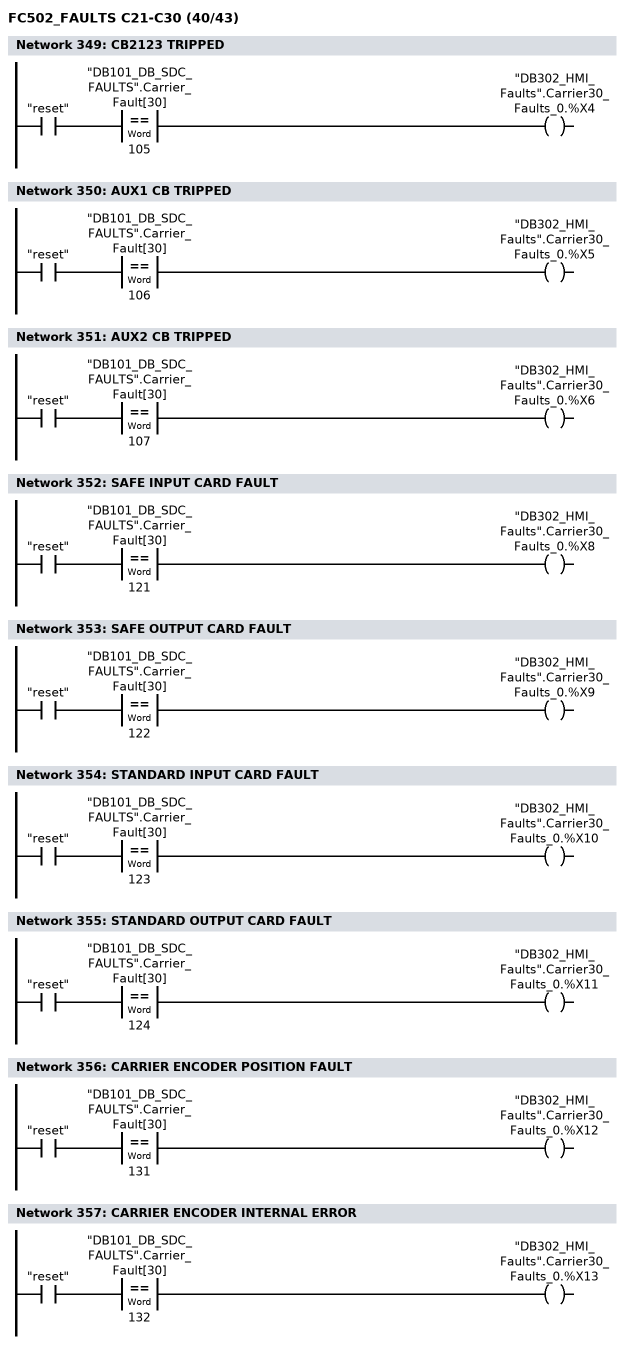
   RUNG wire#powerrail
      Contact( "reset" )
      { S7_Templates := "SrcType := Word" } EQ_Contact(in1 := "DB101_DB_SDC_FAULTS".Carrier_Fault[30], in2 := 105)
      Coil( "DB302_HMI_Faults".Carrier30_Faults_0.%X4 )
   END_RUNG
   // the same network as SCL:
   "DB302_HMI_Faults".Carrier30_Faults_0.%X4 := "reset" AND ("DB101_DB_SDC_FAULTS".Carrier_Fault[30] = 105);
END_REGION

REGION Network 350: AUX1 CB TRIPPED
   RUNG wire#powerrail
      Contact( "reset" )
      { S7_Templates := "SrcType := Word" } EQ_Contact(in1 := "DB101_DB_SDC_FAULTS".Carrier_Fault[30], in2 := 106)
      Coil( "DB302_HMI_Faults".Carrier30_Faults_0.%X5 )
   END_RUNG
   // the same network as SCL:
   "DB302_HMI_Faults".Carrier30_Faults_0.%X5 := "reset" AND ("DB101_DB_SDC_FAULTS".Carrier_Fault[30] = 106);
END_REGION

REGION Network 351: AUX2 CB TRIPPED
   RUNG wire#powerrail
      Contact( "reset" )
      { S7_Templates := "SrcType := Word" } EQ_Contact(in1 := "DB101_DB_SDC_FAULTS".Carrier_Fault[30], in2 := 107)
      Coil( "DB302_HMI_Faults".Carrier30_Faults_0.%X6 )
   END_RUNG
   // the same network as SCL:
   "DB302_HMI_Faults".Carrier30_Faults_0.%X6 := "reset" AND ("DB101_DB_SDC_FAULTS".Carrier_Fault[30] = 107);
END_REGION

REGION Network 352: SAFE INPUT CARD FAULT
   RUNG wire#powerrail
      Contact( "reset" )
      { S7_Templates := "SrcType := Word" } EQ_Contact(in1 := "DB101_DB_SDC_FAULTS".Carrier_Fault[30], in2 := 121)
      Coil( "DB302_HMI_Faults".Carrier30_Faults_0.%X8 )
   END_RUNG
   // the same network as SCL:
   "DB302_HMI_Faults".Carrier30_Faults_0.%X8 := "reset" AND ("DB101_DB_SDC_FAULTS".Carrier_Fault[30] = 121);
END_REGION

REGION Network 353: SAFE OUTPUT CARD FAULT
   RUNG wire#powerrail
      Contact( "reset" )
      { S7_Templates := "SrcType := Word" } EQ_Contact(in1 := "DB101_DB_SDC_FAULTS".Carrier_Fault[30], in2 := 122)
      Coil( "DB302_HMI_Faults".Carrier30_Faults_0.%X9 )
   END_RUNG
   // the same network as SCL:
   "DB302_HMI_Faults".Carrier30_Faults_0.%X9 := "reset" AND ("DB101_DB_SDC_FAULTS".Carrier_Fault[30] = 122);
END_REGION

REGION Network 354: STANDARD INPUT CARD FAULT
   RUNG wire#powerrail
      Contact( "reset" )
      { S7_Templates := "SrcType := Word" } EQ_Contact(in1 := "DB101_DB_SDC_FAULTS".Carrier_Fault[30], in2 := 123)
      Coil( "DB302_HMI_Faults".Carrier30_Faults_0.%X10 )
   END_RUNG
   // the same network as SCL:
   "DB302_HMI_Faults".Carrier30_Faults_0.%X10 := "reset" AND ("DB101_DB_SDC_FAULTS".Carrier_Fault[30] = 123);
END_REGION

REGION Network 355: STANDARD OUTPUT CARD FAULT
   RUNG wire#powerrail
      Contact( "reset" )
      { S7_Templates := "SrcType := Word" } EQ_Contact(in1 := "DB101_DB_SDC_FAULTS".Carrier_Fault[30], in2 := 124)
      Coil( "DB302_HMI_Faults".Carrier30_Faults_0.%X11 )
   END_RUNG
   // the same network as SCL:
   "DB302_HMI_Faults".Carrier30_Faults_0.%X11 := "reset" AND ("DB101_DB_SDC_FAULTS".Carrier_Fault[30] = 124);
END_REGION

REGION Network 356: CARRIER ENCODER POSITION FAULT
   RUNG wire#powerrail
      Contact( "reset" )
      { S7_Templates := "SrcType := Word" } EQ_Contact(in1 := "DB101_DB_SDC_FAULTS".Carrier_Fault[30], in2 := 131)
      Coil( "DB302_HMI_Faults".Carrier30_Faults_0.%X12 )
   END_RUNG
   // the same network as SCL:
   "DB302_HMI_Faults".Carrier30_Faults_0.%X12 := "reset" AND ("DB101_DB_SDC_FAULTS".Carrier_Fault[30] = 131);
END_REGION

REGION Network 357: CARRIER ENCODER INTERNAL ERROR
   RUNG wire#powerrail
      Contact( "reset" )
      { S7_Templates := "SrcType := Word" } EQ_Contact(in1 := "DB101_DB_SDC_FAULTS".Carrier_Fault[30], in2 := 132)
      Coil( "DB302_HMI_Faults".Carrier30_Faults_0.%X13 )
   END_RUNG
   // the same network as SCL:
   "DB302_HMI_Faults".Carrier30_Faults_0.%X13 := "reset" AND ("DB101_DB_SDC_FAULTS".Carrier_Fault[30] = 132);
END_REGION

REGION Network 358: CARRIER ENCODER COMM FAULT
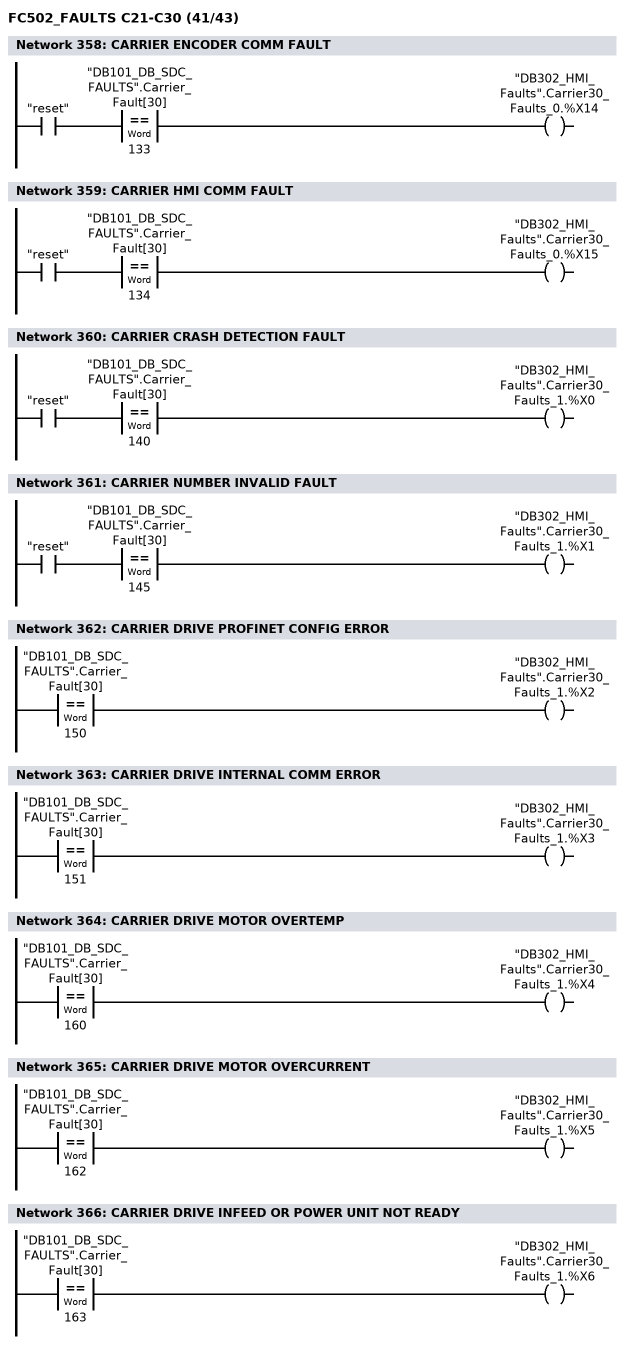
   RUNG wire#powerrail
      Contact( "reset" )
      { S7_Templates := "SrcType := Word" } EQ_Contact(in1 := "DB101_DB_SDC_FAULTS".Carrier_Fault[30], in2 := 133)
      Coil( "DB302_HMI_Faults".Carrier30_Faults_0.%X14 )
   END_RUNG
   // the same network as SCL:
   "DB302_HMI_Faults".Carrier30_Faults_0.%X14 := "reset" AND ("DB101_DB_SDC_FAULTS".Carrier_Fault[30] = 133);
END_REGION

REGION Network 359: CARRIER HMI COMM FAULT
   RUNG wire#powerrail
      Contact( "reset" )
      { S7_Templates := "SrcType := Word" } EQ_Contact(in1 := "DB101_DB_SDC_FAULTS".Carrier_Fault[30], in2 := 134)
      Coil( "DB302_HMI_Faults".Carrier30_Faults_0.%X15 )
   END_RUNG
   // the same network as SCL:
   "DB302_HMI_Faults".Carrier30_Faults_0.%X15 := "reset" AND ("DB101_DB_SDC_FAULTS".Carrier_Fault[30] = 134);
END_REGION

REGION Network 360: CARRIER CRASH DETECTION FAULT
   RUNG wire#powerrail
      Contact( "reset" )
      { S7_Templates := "SrcType := Word" } EQ_Contact(in1 := "DB101_DB_SDC_FAULTS".Carrier_Fault[30], in2 := 140)
      Coil( "DB302_HMI_Faults".Carrier30_Faults_1.%X0 )
   END_RUNG
   // the same network as SCL:
   "DB302_HMI_Faults".Carrier30_Faults_1.%X0 := "reset" AND ("DB101_DB_SDC_FAULTS".Carrier_Fault[30] = 140);
END_REGION

REGION Network 361: CARRIER NUMBER INVALID FAULT
   RUNG wire#powerrail
      Contact( "reset" )
      { S7_Templates := "SrcType := Word" } EQ_Contact(in1 := "DB101_DB_SDC_FAULTS".Carrier_Fault[30], in2 := 145)
      Coil( "DB302_HMI_Faults".Carrier30_Faults_1.%X1 )
   END_RUNG
   // the same network as SCL:
   "DB302_HMI_Faults".Carrier30_Faults_1.%X1 := "reset" AND ("DB101_DB_SDC_FAULTS".Carrier_Fault[30] = 145);
END_REGION

REGION Network 362: CARRIER DRIVE PROFINET CONFIG ERROR
   RUNG wire#powerrail
      { S7_Templates := "SrcType := Word" } EQ_Contact(in1 := "DB101_DB_SDC_FAULTS".Carrier_Fault[30], in2 := 150)
      Coil( "DB302_HMI_Faults".Carrier30_Faults_1.%X2 )
   END_RUNG
   // the same network as SCL:
   "DB302_HMI_Faults".Carrier30_Faults_1.%X2 := "DB101_DB_SDC_FAULTS".Carrier_Fault[30] = 150;
END_REGION

REGION Network 363: CARRIER DRIVE INTERNAL COMM ERROR
   RUNG wire#powerrail
      { S7_Templates := "SrcType := Word" } EQ_Contact(in1 := "DB101_DB_SDC_FAULTS".Carrier_Fault[30], in2 := 151)
      Coil( "DB302_HMI_Faults".Carrier30_Faults_1.%X3 )
   END_RUNG
   // the same network as SCL:
   "DB302_HMI_Faults".Carrier30_Faults_1.%X3 := "DB101_DB_SDC_FAULTS".Carrier_Fault[30] = 151;
END_REGION

REGION Network 364: CARRIER DRIVE MOTOR OVERTEMP
   RUNG wire#powerrail
      { S7_Templates := "SrcType := Word" } EQ_Contact(in1 := "DB101_DB_SDC_FAULTS".Carrier_Fault[30], in2 := 160)
      Coil( "DB302_HMI_Faults".Carrier30_Faults_1.%X4 )
   END_RUNG
   // the same network as SCL:
   "DB302_HMI_Faults".Carrier30_Faults_1.%X4 := "DB101_DB_SDC_FAULTS".Carrier_Fault[30] = 160;
END_REGION

REGION Network 365: CARRIER DRIVE MOTOR OVERCURRENT
   RUNG wire#powerrail
      { S7_Templates := "SrcType := Word" } EQ_Contact(in1 := "DB101_DB_SDC_FAULTS".Carrier_Fault[30], in2 := 162)
      Coil( "DB302_HMI_Faults".Carrier30_Faults_1.%X5 )
   END_RUNG
   // the same network as SCL:
   "DB302_HMI_Faults".Carrier30_Faults_1.%X5 := "DB101_DB_SDC_FAULTS".Carrier_Fault[30] = 162;
END_REGION

REGION Network 366: CARRIER DRIVE INFEED OR POWER UNIT NOT READY
   RUNG wire#powerrail
      { S7_Templates := "SrcType := Word" } EQ_Contact(in1 := "DB101_DB_SDC_FAULTS".Carrier_Fault[30], in2 := 163)
      Coil( "DB302_HMI_Faults".Carrier30_Faults_1.%X6 )
   END_RUNG
   // the same network as SCL:
   "DB302_HMI_Faults".Carrier30_Faults_1.%X6 := "DB101_DB_SDC_FAULTS".Carrier_Fault[30] = 163;
END_REGION

REGION Network 367: CARRIER DRIVE SHORT CIRCUIT / GROUND FAULT DETECTED
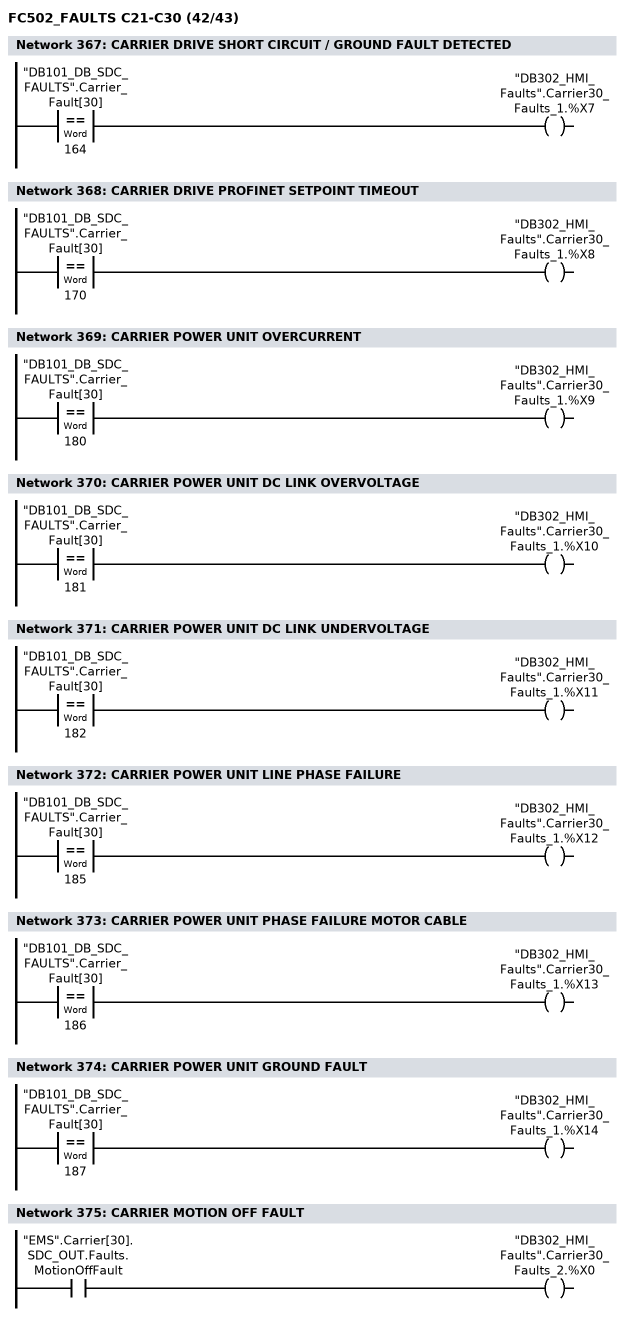
   RUNG wire#powerrail
      { S7_Templates := "SrcType := Word" } EQ_Contact(in1 := "DB101_DB_SDC_FAULTS".Carrier_Fault[30], in2 := 164)
      Coil( "DB302_HMI_Faults".Carrier30_Faults_1.%X7 )
   END_RUNG
   // the same network as SCL:
   "DB302_HMI_Faults".Carrier30_Faults_1.%X7 := "DB101_DB_SDC_FAULTS".Carrier_Fault[30] = 164;
END_REGION

REGION Network 368: CARRIER DRIVE PROFINET SETPOINT TIMEOUT
   RUNG wire#powerrail
      { S7_Templates := "SrcType := Word" } EQ_Contact(in1 := "DB101_DB_SDC_FAULTS".Carrier_Fault[30], in2 := 170)
      Coil( "DB302_HMI_Faults".Carrier30_Faults_1.%X8 )
   END_RUNG
   // the same network as SCL:
   "DB302_HMI_Faults".Carrier30_Faults_1.%X8 := "DB101_DB_SDC_FAULTS".Carrier_Fault[30] = 170;
END_REGION

REGION Network 369: CARRIER POWER UNIT OVERCURRENT
   RUNG wire#powerrail
      { S7_Templates := "SrcType := Word" } EQ_Contact(in1 := "DB101_DB_SDC_FAULTS".Carrier_Fault[30], in2 := 180)
      Coil( "DB302_HMI_Faults".Carrier30_Faults_1.%X9 )
   END_RUNG
   // the same network as SCL:
   "DB302_HMI_Faults".Carrier30_Faults_1.%X9 := "DB101_DB_SDC_FAULTS".Carrier_Fault[30] = 180;
END_REGION

REGION Network 370: CARRIER POWER UNIT DC LINK OVERVOLTAGE
   RUNG wire#powerrail
      { S7_Templates := "SrcType := Word" } EQ_Contact(in1 := "DB101_DB_SDC_FAULTS".Carrier_Fault[30], in2 := 181)
      Coil( "DB302_HMI_Faults".Carrier30_Faults_1.%X10 )
   END_RUNG
   // the same network as SCL:
   "DB302_HMI_Faults".Carrier30_Faults_1.%X10 := "DB101_DB_SDC_FAULTS".Carrier_Fault[30] = 181;
END_REGION

REGION Network 371: CARRIER POWER UNIT DC LINK UNDERVOLTAGE
   RUNG wire#powerrail
      { S7_Templates := "SrcType := Word" } EQ_Contact(in1 := "DB101_DB_SDC_FAULTS".Carrier_Fault[30], in2 := 182)
      Coil( "DB302_HMI_Faults".Carrier30_Faults_1.%X11 )
   END_RUNG
   // the same network as SCL:
   "DB302_HMI_Faults".Carrier30_Faults_1.%X11 := "DB101_DB_SDC_FAULTS".Carrier_Fault[30] = 182;
END_REGION

REGION Network 372: CARRIER POWER UNIT LINE PHASE FAILURE
   RUNG wire#powerrail
      { S7_Templates := "SrcType := Word" } EQ_Contact(in1 := "DB101_DB_SDC_FAULTS".Carrier_Fault[30], in2 := 185)
      Coil( "DB302_HMI_Faults".Carrier30_Faults_1.%X12 )
   END_RUNG
   // the same network as SCL:
   "DB302_HMI_Faults".Carrier30_Faults_1.%X12 := "DB101_DB_SDC_FAULTS".Carrier_Fault[30] = 185;
END_REGION

REGION Network 373: CARRIER POWER UNIT PHASE FAILURE MOTOR CABLE
   RUNG wire#powerrail
      { S7_Templates := "SrcType := Word" } EQ_Contact(in1 := "DB101_DB_SDC_FAULTS".Carrier_Fault[30], in2 := 186)
      Coil( "DB302_HMI_Faults".Carrier30_Faults_1.%X13 )
   END_RUNG
   // the same network as SCL:
   "DB302_HMI_Faults".Carrier30_Faults_1.%X13 := "DB101_DB_SDC_FAULTS".Carrier_Fault[30] = 186;
END_REGION

REGION Network 374: CARRIER POWER UNIT GROUND FAULT
   RUNG wire#powerrail
      { S7_Templates := "SrcType := Word" } EQ_Contact(in1 := "DB101_DB_SDC_FAULTS".Carrier_Fault[30], in2 := 187)
      Coil( "DB302_HMI_Faults".Carrier30_Faults_1.%X14 )
   END_RUNG
   // the same network as SCL:
   "DB302_HMI_Faults".Carrier30_Faults_1.%X14 := "DB101_DB_SDC_FAULTS".Carrier_Fault[30] = 187;
END_REGION

REGION Network 375: CARRIER MOTION OFF FAULT
   RUNG wire#powerrail
      Contact( "EMS".Carrier[30].SDC_OUT.Faults.MotionOffFault )
      Coil( "DB302_HMI_Faults".Carrier30_Faults_2.%X0 )
   END_RUNG
   // the same network as SCL:
   "DB302_HMI_Faults".Carrier30_Faults_2.%X0 := "EMS".Carrier[30].SDC_OUT.Faults.MotionOffFault;
END_REGION

REGION Network 376: CARRIER MOTION ON FAULT
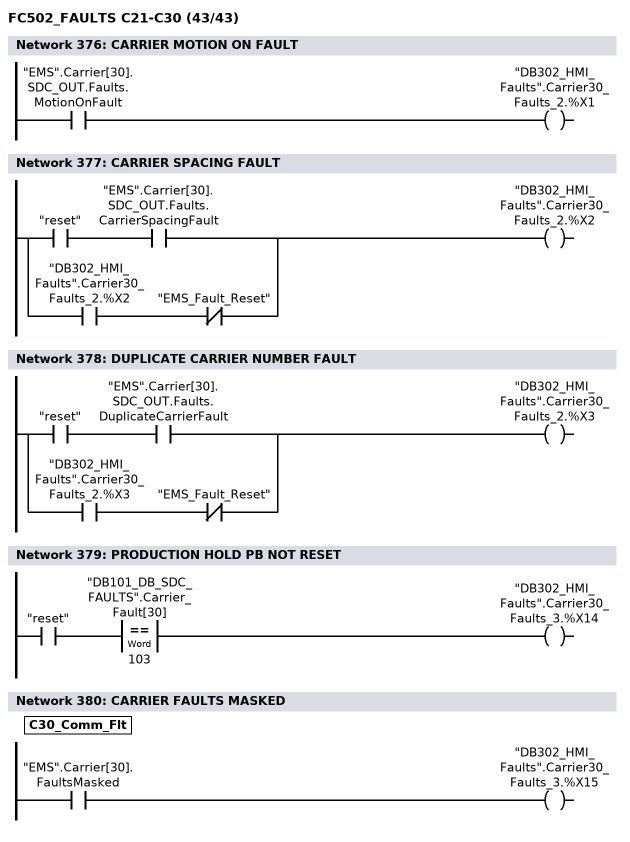
   RUNG wire#powerrail
      Contact( "EMS".Carrier[30].SDC_OUT.Faults.MotionOnFault )
      Coil( "DB302_HMI_Faults".Carrier30_Faults_2.%X1 )
   END_RUNG
   // the same network as SCL:
   "DB302_HMI_Faults".Carrier30_Faults_2.%X1 := "EMS".Carrier[30].SDC_OUT.Faults.MotionOnFault;
END_REGION

REGION Network 377: CARRIER SPACING FAULT
   RUNG wire#powerrail
      Contact( "reset" )
      Contact( "EMS".Carrier[30].SDC_OUT.Faults.CarrierSpacingFault )
      wire#w1
      Coil( "DB302_HMI_Faults".Carrier30_Faults_2.%X2 )
   END_RUNG
   RUNG wire#powerrail
      Contact( "DB302_HMI_Faults".Carrier30_Faults_2.%X2 )
      I_Contact( "EMS_Fault_Reset" )
   END_RUNG wire#w1
   // the same network as SCL:
   "DB302_HMI_Faults".Carrier30_Faults_2.%X2 := ("reset" AND "EMS".Carrier[30].SDC_OUT.Faults.CarrierSpacingFault) OR ("DB302_HMI_Faults".Carrier30_Faults_2.%X2 AND NOT "EMS_Fault_Reset");
END_REGION

REGION Network 378: DUPLICATE CARRIER NUMBER FAULT
   RUNG wire#powerrail
      Contact( "reset" )
      Contact( "EMS".Carrier[30].SDC_OUT.Faults.DuplicateCarrierFault )
      wire#w1
      Coil( "DB302_HMI_Faults".Carrier30_Faults_2.%X3 )
   END_RUNG
   RUNG wire#powerrail
      Contact( "DB302_HMI_Faults".Carrier30_Faults_2.%X3 )
      I_Contact( "EMS_Fault_Reset" )
   END_RUNG wire#w1
   // the same network as SCL:
   "DB302_HMI_Faults".Carrier30_Faults_2.%X3 := ("reset" AND "EMS".Carrier[30].SDC_OUT.Faults.DuplicateCarrierFault) OR ("DB302_HMI_Faults".Carrier30_Faults_2.%X3 AND NOT "EMS_Fault_Reset");
END_REGION

REGION Network 379: PRODUCTION HOLD PB NOT RESET
   RUNG wire#powerrail
      Contact( "reset" )
      { S7_Templates := "SrcType := Word" } EQ_Contact(in1 := "DB101_DB_SDC_FAULTS".Carrier_Fault[30], in2 := 103)
      Coil( "DB302_HMI_Faults".Carrier30_Faults_3.%X14 )
   END_RUNG
   // the same network as SCL:
   "DB302_HMI_Faults".Carrier30_Faults_3.%X14 := "reset" AND ("DB101_DB_SDC_FAULTS".Carrier_Fault[30] = 103);
END_REGION

REGION Network 380: CARRIER FAULTS MASKED
   Label( C30_Comm_Flt )
   RUNG wire#powerrail
      Contact( "EMS".Carrier[30].FaultsMasked )
      Coil( "DB302_HMI_Faults".Carrier30_Faults_3.%X15 )
   END_RUNG
   // the same network as SCL:
   C30_Comm_Flt:
   "DB302_HMI_Faults".Carrier30_Faults_3.%X15 := "EMS".Carrier[30].FaultsMasked;
END_REGION
END_FUNCTION

FUNCTION "FC503_FAULTS C31-C40" : Void   // FC503, LAD
{ S7_Optimized_Access := 'TRUE' }
VERSION : 0.1
BEGIN

REGION Network 1: CARRIER 31 FAULTS
END_REGION

REGION Network 2: CARRIER PLC NOT COMMUNICATING
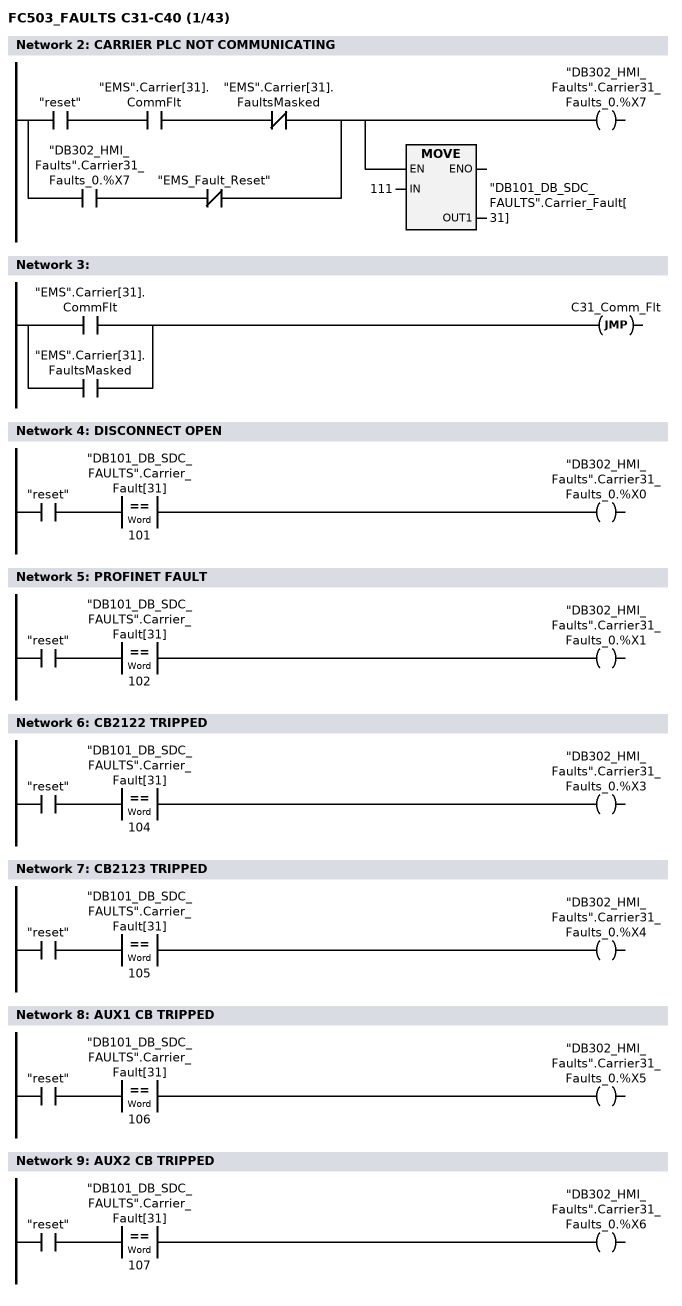
   RUNG wire#powerrail
      Contact( "reset" )
      Contact( "EMS".Carrier[31].CommFlt )
      I_Contact( "EMS".Carrier[31].FaultsMasked )
      wire#w1
      Coil( "DB302_HMI_Faults".Carrier31_Faults_0.%X7 )
   END_RUNG
   RUNG wire#powerrail
      Contact( "DB302_HMI_Faults".Carrier31_Faults_0.%X7 )
      I_Contact( "EMS_Fault_Reset" )
   END_RUNG wire#w1
   RUNG wire#w1
      Move(in := 111, out1 => "DB101_DB_SDC_FAULTS".Carrier_Fault[31])
   END_RUNG
   // the same network as SCL:
   "DB302_HMI_Faults".Carrier31_Faults_0.%X7 := ("reset" AND "EMS".Carrier[31].CommFlt AND NOT "EMS".Carrier[31].FaultsMasked) OR ("DB302_HMI_Faults".Carrier31_Faults_0.%X7 AND NOT "EMS_Fault_Reset");
   IF "DB302_HMI_Faults".Carrier31_Faults_0.%X7 THEN "DB101_DB_SDC_FAULTS".Carrier_Fault[31] := 111; END_IF;
END_REGION

REGION Network 3
   RUNG wire#powerrail
      Contact( "EMS".Carrier[31].CommFlt )
      wire#w1
      JumpCoil( C31_Comm_Flt )
   END_RUNG
   RUNG wire#powerrail
      Contact( "EMS".Carrier[31].FaultsMasked )
   END_RUNG wire#w1
   // the same network as SCL:
   IF "EMS".Carrier[31].CommFlt OR "EMS".Carrier[31].FaultsMasked THEN GOTO C31_Comm_Flt; END_IF;
END_REGION

REGION Network 4: DISCONNECT OPEN
   RUNG wire#powerrail
      Contact( "reset" )
      { S7_Templates := "SrcType := Word" } EQ_Contact(in1 := "DB101_DB_SDC_FAULTS".Carrier_Fault[31], in2 := 101)
      Coil( "DB302_HMI_Faults".Carrier31_Faults_0.%X0 )
   END_RUNG
   // the same network as SCL:
   "DB302_HMI_Faults".Carrier31_Faults_0.%X0 := "reset" AND ("DB101_DB_SDC_FAULTS".Carrier_Fault[31] = 101);
END_REGION

REGION Network 5: PROFINET FAULT
   RUNG wire#powerrail
      Contact( "reset" )
      { S7_Templates := "SrcType := Word" } EQ_Contact(in1 := "DB101_DB_SDC_FAULTS".Carrier_Fault[31], in2 := 102)
      Coil( "DB302_HMI_Faults".Carrier31_Faults_0.%X1 )
   END_RUNG
   // the same network as SCL:
   "DB302_HMI_Faults".Carrier31_Faults_0.%X1 := "reset" AND ("DB101_DB_SDC_FAULTS".Carrier_Fault[31] = 102);
END_REGION

REGION Network 6: CB2122 TRIPPED
   RUNG wire#powerrail
      Contact( "reset" )
      { S7_Templates := "SrcType := Word" } EQ_Contact(in1 := "DB101_DB_SDC_FAULTS".Carrier_Fault[31], in2 := 104)
      Coil( "DB302_HMI_Faults".Carrier31_Faults_0.%X3 )
   END_RUNG
   // the same network as SCL:
   "DB302_HMI_Faults".Carrier31_Faults_0.%X3 := "reset" AND ("DB101_DB_SDC_FAULTS".Carrier_Fault[31] = 104);
END_REGION

REGION Network 7: CB2123 TRIPPED
   RUNG wire#powerrail
      Contact( "reset" )
      { S7_Templates := "SrcType := Word" } EQ_Contact(in1 := "DB101_DB_SDC_FAULTS".Carrier_Fault[31], in2 := 105)
      Coil( "DB302_HMI_Faults".Carrier31_Faults_0.%X4 )
   END_RUNG
   // the same network as SCL:
   "DB302_HMI_Faults".Carrier31_Faults_0.%X4 := "reset" AND ("DB101_DB_SDC_FAULTS".Carrier_Fault[31] = 105);
END_REGION

REGION Network 8: AUX1 CB TRIPPED
   RUNG wire#powerrail
      Contact( "reset" )
      { S7_Templates := "SrcType := Word" } EQ_Contact(in1 := "DB101_DB_SDC_FAULTS".Carrier_Fault[31], in2 := 106)
      Coil( "DB302_HMI_Faults".Carrier31_Faults_0.%X5 )
   END_RUNG
   // the same network as SCL:
   "DB302_HMI_Faults".Carrier31_Faults_0.%X5 := "reset" AND ("DB101_DB_SDC_FAULTS".Carrier_Fault[31] = 106);
END_REGION

REGION Network 9: AUX2 CB TRIPPED
   RUNG wire#powerrail
      Contact( "reset" )
      { S7_Templates := "SrcType := Word" } EQ_Contact(in1 := "DB101_DB_SDC_FAULTS".Carrier_Fault[31], in2 := 107)
      Coil( "DB302_HMI_Faults".Carrier31_Faults_0.%X6 )
   END_RUNG
   // the same network as SCL:
   "DB302_HMI_Faults".Carrier31_Faults_0.%X6 := "reset" AND ("DB101_DB_SDC_FAULTS".Carrier_Fault[31] = 107);
END_REGION

REGION Network 10: SAFE INPUT CARD FAULT
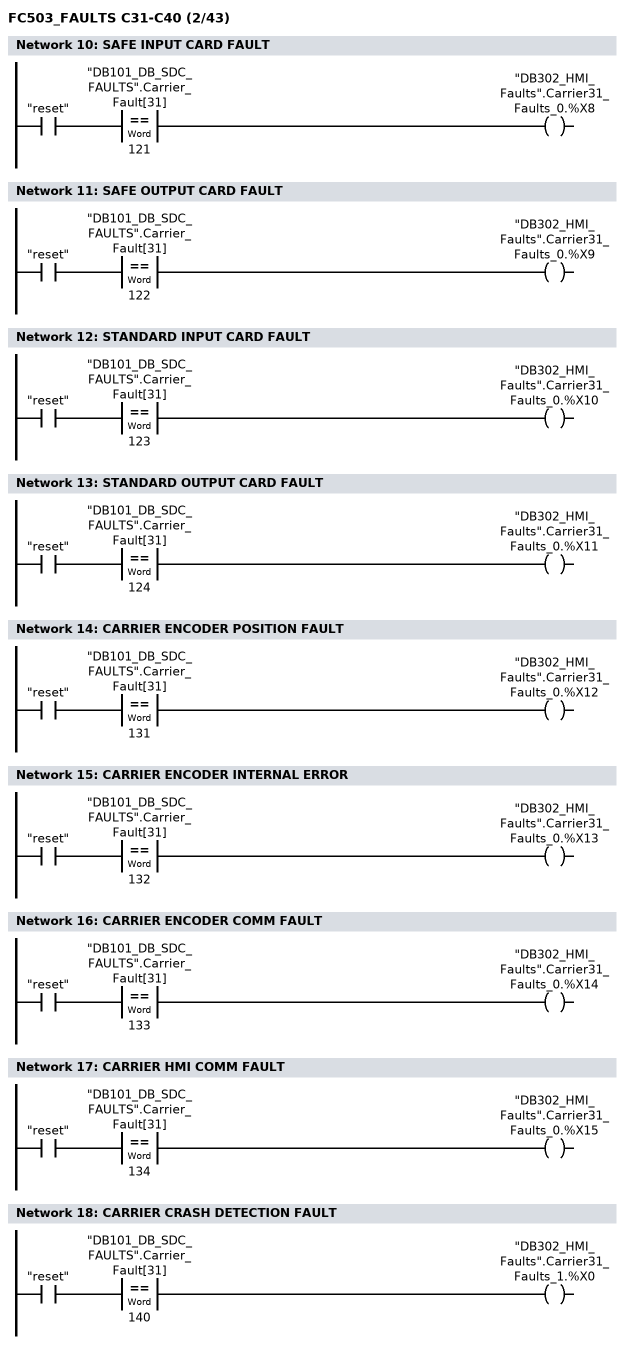
   RUNG wire#powerrail
      Contact( "reset" )
      { S7_Templates := "SrcType := Word" } EQ_Contact(in1 := "DB101_DB_SDC_FAULTS".Carrier_Fault[31], in2 := 121)
      Coil( "DB302_HMI_Faults".Carrier31_Faults_0.%X8 )
   END_RUNG
   // the same network as SCL:
   "DB302_HMI_Faults".Carrier31_Faults_0.%X8 := "reset" AND ("DB101_DB_SDC_FAULTS".Carrier_Fault[31] = 121);
END_REGION

REGION Network 11: SAFE OUTPUT CARD FAULT
   RUNG wire#powerrail
      Contact( "reset" )
      { S7_Templates := "SrcType := Word" } EQ_Contact(in1 := "DB101_DB_SDC_FAULTS".Carrier_Fault[31], in2 := 122)
      Coil( "DB302_HMI_Faults".Carrier31_Faults_0.%X9 )
   END_RUNG
   // the same network as SCL:
   "DB302_HMI_Faults".Carrier31_Faults_0.%X9 := "reset" AND ("DB101_DB_SDC_FAULTS".Carrier_Fault[31] = 122);
END_REGION

REGION Network 12: STANDARD INPUT CARD FAULT
   RUNG wire#powerrail
      Contact( "reset" )
      { S7_Templates := "SrcType := Word" } EQ_Contact(in1 := "DB101_DB_SDC_FAULTS".Carrier_Fault[31], in2 := 123)
      Coil( "DB302_HMI_Faults".Carrier31_Faults_0.%X10 )
   END_RUNG
   // the same network as SCL:
   "DB302_HMI_Faults".Carrier31_Faults_0.%X10 := "reset" AND ("DB101_DB_SDC_FAULTS".Carrier_Fault[31] = 123);
END_REGION

REGION Network 13: STANDARD OUTPUT CARD FAULT
   RUNG wire#powerrail
      Contact( "reset" )
      { S7_Templates := "SrcType := Word" } EQ_Contact(in1 := "DB101_DB_SDC_FAULTS".Carrier_Fault[31], in2 := 124)
      Coil( "DB302_HMI_Faults".Carrier31_Faults_0.%X11 )
   END_RUNG
   // the same network as SCL:
   "DB302_HMI_Faults".Carrier31_Faults_0.%X11 := "reset" AND ("DB101_DB_SDC_FAULTS".Carrier_Fault[31] = 124);
END_REGION

REGION Network 14: CARRIER ENCODER POSITION FAULT
   RUNG wire#powerrail
      Contact( "reset" )
      { S7_Templates := "SrcType := Word" } EQ_Contact(in1 := "DB101_DB_SDC_FAULTS".Carrier_Fault[31], in2 := 131)
      Coil( "DB302_HMI_Faults".Carrier31_Faults_0.%X12 )
   END_RUNG
   // the same network as SCL:
   "DB302_HMI_Faults".Carrier31_Faults_0.%X12 := "reset" AND ("DB101_DB_SDC_FAULTS".Carrier_Fault[31] = 131);
END_REGION

REGION Network 15: CARRIER ENCODER INTERNAL ERROR
   RUNG wire#powerrail
      Contact( "reset" )
      { S7_Templates := "SrcType := Word" } EQ_Contact(in1 := "DB101_DB_SDC_FAULTS".Carrier_Fault[31], in2 := 132)
      Coil( "DB302_HMI_Faults".Carrier31_Faults_0.%X13 )
   END_RUNG
   // the same network as SCL:
   "DB302_HMI_Faults".Carrier31_Faults_0.%X13 := "reset" AND ("DB101_DB_SDC_FAULTS".Carrier_Fault[31] = 132);
END_REGION

REGION Network 16: CARRIER ENCODER COMM FAULT
   RUNG wire#powerrail
      Contact( "reset" )
      { S7_Templates := "SrcType := Word" } EQ_Contact(in1 := "DB101_DB_SDC_FAULTS".Carrier_Fault[31], in2 := 133)
      Coil( "DB302_HMI_Faults".Carrier31_Faults_0.%X14 )
   END_RUNG
   // the same network as SCL:
   "DB302_HMI_Faults".Carrier31_Faults_0.%X14 := "reset" AND ("DB101_DB_SDC_FAULTS".Carrier_Fault[31] = 133);
END_REGION

REGION Network 17: CARRIER HMI COMM FAULT
   RUNG wire#powerrail
      Contact( "reset" )
      { S7_Templates := "SrcType := Word" } EQ_Contact(in1 := "DB101_DB_SDC_FAULTS".Carrier_Fault[31], in2 := 134)
      Coil( "DB302_HMI_Faults".Carrier31_Faults_0.%X15 )
   END_RUNG
   // the same network as SCL:
   "DB302_HMI_Faults".Carrier31_Faults_0.%X15 := "reset" AND ("DB101_DB_SDC_FAULTS".Carrier_Fault[31] = 134);
END_REGION

REGION Network 18: CARRIER CRASH DETECTION FAULT
   RUNG wire#powerrail
      Contact( "reset" )
      { S7_Templates := "SrcType := Word" } EQ_Contact(in1 := "DB101_DB_SDC_FAULTS".Carrier_Fault[31], in2 := 140)
      Coil( "DB302_HMI_Faults".Carrier31_Faults_1.%X0 )
   END_RUNG
   // the same network as SCL:
   "DB302_HMI_Faults".Carrier31_Faults_1.%X0 := "reset" AND ("DB101_DB_SDC_FAULTS".Carrier_Fault[31] = 140);
END_REGION

REGION Network 19: CARRIER NUMBER INVALID FAULT
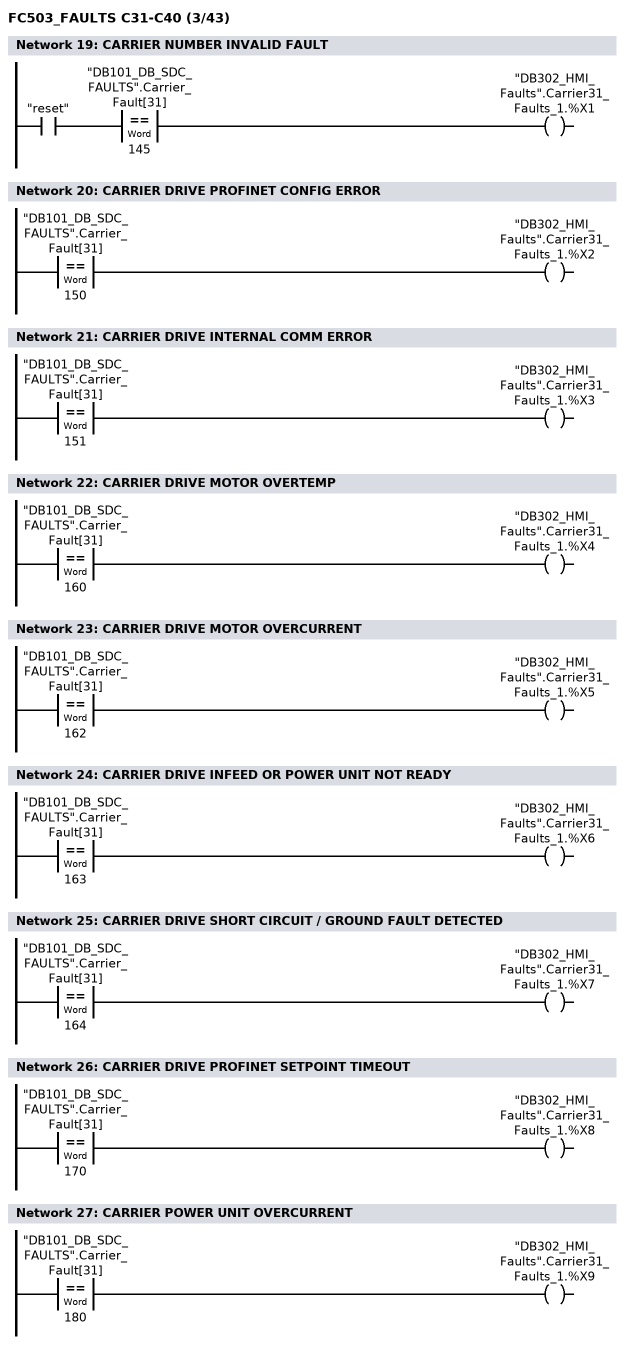
   RUNG wire#powerrail
      Contact( "reset" )
      { S7_Templates := "SrcType := Word" } EQ_Contact(in1 := "DB101_DB_SDC_FAULTS".Carrier_Fault[31], in2 := 145)
      Coil( "DB302_HMI_Faults".Carrier31_Faults_1.%X1 )
   END_RUNG
   // the same network as SCL:
   "DB302_HMI_Faults".Carrier31_Faults_1.%X1 := "reset" AND ("DB101_DB_SDC_FAULTS".Carrier_Fault[31] = 145);
END_REGION

REGION Network 20: CARRIER DRIVE PROFINET CONFIG ERROR
   RUNG wire#powerrail
      { S7_Templates := "SrcType := Word" } EQ_Contact(in1 := "DB101_DB_SDC_FAULTS".Carrier_Fault[31], in2 := 150)
      Coil( "DB302_HMI_Faults".Carrier31_Faults_1.%X2 )
   END_RUNG
   // the same network as SCL:
   "DB302_HMI_Faults".Carrier31_Faults_1.%X2 := "DB101_DB_SDC_FAULTS".Carrier_Fault[31] = 150;
END_REGION

REGION Network 21: CARRIER DRIVE INTERNAL COMM ERROR
   RUNG wire#powerrail
      { S7_Templates := "SrcType := Word" } EQ_Contact(in1 := "DB101_DB_SDC_FAULTS".Carrier_Fault[31], in2 := 151)
      Coil( "DB302_HMI_Faults".Carrier31_Faults_1.%X3 )
   END_RUNG
   // the same network as SCL:
   "DB302_HMI_Faults".Carrier31_Faults_1.%X3 := "DB101_DB_SDC_FAULTS".Carrier_Fault[31] = 151;
END_REGION

REGION Network 22: CARRIER DRIVE MOTOR OVERTEMP
   RUNG wire#powerrail
      { S7_Templates := "SrcType := Word" } EQ_Contact(in1 := "DB101_DB_SDC_FAULTS".Carrier_Fault[31], in2 := 160)
      Coil( "DB302_HMI_Faults".Carrier31_Faults_1.%X4 )
   END_RUNG
   // the same network as SCL:
   "DB302_HMI_Faults".Carrier31_Faults_1.%X4 := "DB101_DB_SDC_FAULTS".Carrier_Fault[31] = 160;
END_REGION

REGION Network 23: CARRIER DRIVE MOTOR OVERCURRENT
   RUNG wire#powerrail
      { S7_Templates := "SrcType := Word" } EQ_Contact(in1 := "DB101_DB_SDC_FAULTS".Carrier_Fault[31], in2 := 162)
      Coil( "DB302_HMI_Faults".Carrier31_Faults_1.%X5 )
   END_RUNG
   // the same network as SCL:
   "DB302_HMI_Faults".Carrier31_Faults_1.%X5 := "DB101_DB_SDC_FAULTS".Carrier_Fault[31] = 162;
END_REGION

REGION Network 24: CARRIER DRIVE INFEED OR POWER UNIT NOT READY
   RUNG wire#powerrail
      { S7_Templates := "SrcType := Word" } EQ_Contact(in1 := "DB101_DB_SDC_FAULTS".Carrier_Fault[31], in2 := 163)
      Coil( "DB302_HMI_Faults".Carrier31_Faults_1.%X6 )
   END_RUNG
   // the same network as SCL:
   "DB302_HMI_Faults".Carrier31_Faults_1.%X6 := "DB101_DB_SDC_FAULTS".Carrier_Fault[31] = 163;
END_REGION

REGION Network 25: CARRIER DRIVE SHORT CIRCUIT / GROUND FAULT DETECTED
   RUNG wire#powerrail
      { S7_Templates := "SrcType := Word" } EQ_Contact(in1 := "DB101_DB_SDC_FAULTS".Carrier_Fault[31], in2 := 164)
      Coil( "DB302_HMI_Faults".Carrier31_Faults_1.%X7 )
   END_RUNG
   // the same network as SCL:
   "DB302_HMI_Faults".Carrier31_Faults_1.%X7 := "DB101_DB_SDC_FAULTS".Carrier_Fault[31] = 164;
END_REGION

REGION Network 26: CARRIER DRIVE PROFINET SETPOINT TIMEOUT
   RUNG wire#powerrail
      { S7_Templates := "SrcType := Word" } EQ_Contact(in1 := "DB101_DB_SDC_FAULTS".Carrier_Fault[31], in2 := 170)
      Coil( "DB302_HMI_Faults".Carrier31_Faults_1.%X8 )
   END_RUNG
   // the same network as SCL:
   "DB302_HMI_Faults".Carrier31_Faults_1.%X8 := "DB101_DB_SDC_FAULTS".Carrier_Fault[31] = 170;
END_REGION

REGION Network 27: CARRIER POWER UNIT OVERCURRENT
   RUNG wire#powerrail
      { S7_Templates := "SrcType := Word" } EQ_Contact(in1 := "DB101_DB_SDC_FAULTS".Carrier_Fault[31], in2 := 180)
      Coil( "DB302_HMI_Faults".Carrier31_Faults_1.%X9 )
   END_RUNG
   // the same network as SCL:
   "DB302_HMI_Faults".Carrier31_Faults_1.%X9 := "DB101_DB_SDC_FAULTS".Carrier_Fault[31] = 180;
END_REGION

REGION Network 28: CARRIER POWER UNIT DC LINK OVERVOLTAGE
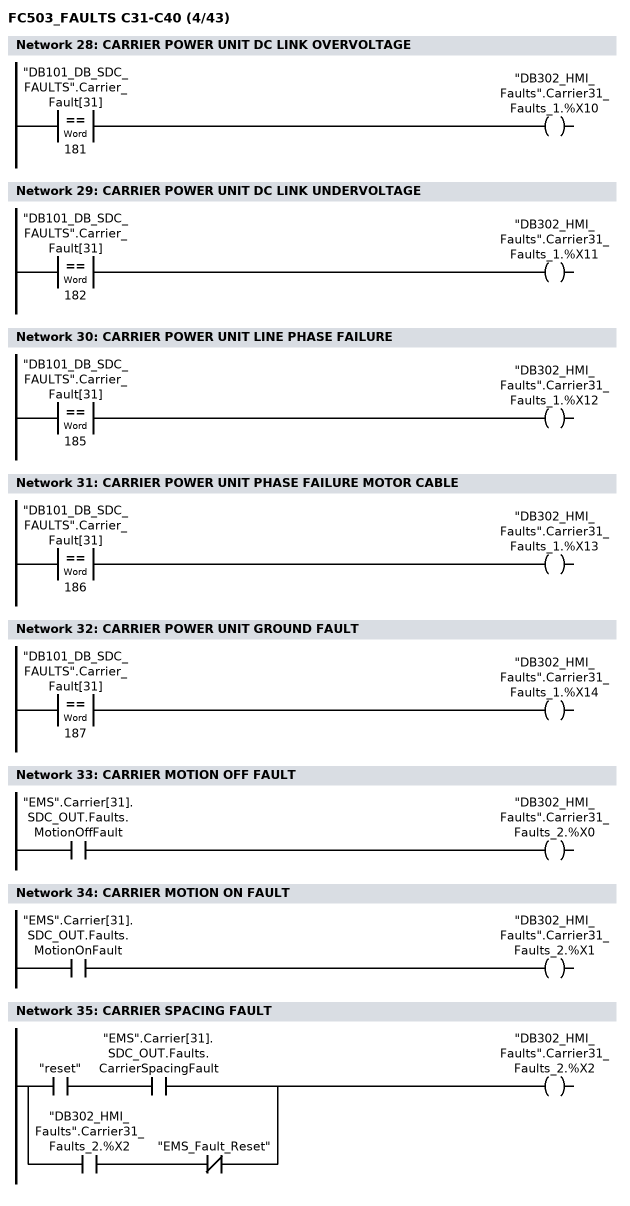
   RUNG wire#powerrail
      { S7_Templates := "SrcType := Word" } EQ_Contact(in1 := "DB101_DB_SDC_FAULTS".Carrier_Fault[31], in2 := 181)
      Coil( "DB302_HMI_Faults".Carrier31_Faults_1.%X10 )
   END_RUNG
   // the same network as SCL:
   "DB302_HMI_Faults".Carrier31_Faults_1.%X10 := "DB101_DB_SDC_FAULTS".Carrier_Fault[31] = 181;
END_REGION

REGION Network 29: CARRIER POWER UNIT DC LINK UNDERVOLTAGE
   RUNG wire#powerrail
      { S7_Templates := "SrcType := Word" } EQ_Contact(in1 := "DB101_DB_SDC_FAULTS".Carrier_Fault[31], in2 := 182)
      Coil( "DB302_HMI_Faults".Carrier31_Faults_1.%X11 )
   END_RUNG
   // the same network as SCL:
   "DB302_HMI_Faults".Carrier31_Faults_1.%X11 := "DB101_DB_SDC_FAULTS".Carrier_Fault[31] = 182;
END_REGION

REGION Network 30: CARRIER POWER UNIT LINE PHASE FAILURE
   RUNG wire#powerrail
      { S7_Templates := "SrcType := Word" } EQ_Contact(in1 := "DB101_DB_SDC_FAULTS".Carrier_Fault[31], in2 := 185)
      Coil( "DB302_HMI_Faults".Carrier31_Faults_1.%X12 )
   END_RUNG
   // the same network as SCL:
   "DB302_HMI_Faults".Carrier31_Faults_1.%X12 := "DB101_DB_SDC_FAULTS".Carrier_Fault[31] = 185;
END_REGION

REGION Network 31: CARRIER POWER UNIT PHASE FAILURE MOTOR CABLE
   RUNG wire#powerrail
      { S7_Templates := "SrcType := Word" } EQ_Contact(in1 := "DB101_DB_SDC_FAULTS".Carrier_Fault[31], in2 := 186)
      Coil( "DB302_HMI_Faults".Carrier31_Faults_1.%X13 )
   END_RUNG
   // the same network as SCL:
   "DB302_HMI_Faults".Carrier31_Faults_1.%X13 := "DB101_DB_SDC_FAULTS".Carrier_Fault[31] = 186;
END_REGION

REGION Network 32: CARRIER POWER UNIT GROUND FAULT
   RUNG wire#powerrail
      { S7_Templates := "SrcType := Word" } EQ_Contact(in1 := "DB101_DB_SDC_FAULTS".Carrier_Fault[31], in2 := 187)
      Coil( "DB302_HMI_Faults".Carrier31_Faults_1.%X14 )
   END_RUNG
   // the same network as SCL:
   "DB302_HMI_Faults".Carrier31_Faults_1.%X14 := "DB101_DB_SDC_FAULTS".Carrier_Fault[31] = 187;
END_REGION

REGION Network 33: CARRIER MOTION OFF FAULT
   RUNG wire#powerrail
      Contact( "EMS".Carrier[31].SDC_OUT.Faults.MotionOffFault )
      Coil( "DB302_HMI_Faults".Carrier31_Faults_2.%X0 )
   END_RUNG
   // the same network as SCL:
   "DB302_HMI_Faults".Carrier31_Faults_2.%X0 := "EMS".Carrier[31].SDC_OUT.Faults.MotionOffFault;
END_REGION

REGION Network 34: CARRIER MOTION ON FAULT
   RUNG wire#powerrail
      Contact( "EMS".Carrier[31].SDC_OUT.Faults.MotionOnFault )
      Coil( "DB302_HMI_Faults".Carrier31_Faults_2.%X1 )
   END_RUNG
   // the same network as SCL:
   "DB302_HMI_Faults".Carrier31_Faults_2.%X1 := "EMS".Carrier[31].SDC_OUT.Faults.MotionOnFault;
END_REGION

REGION Network 35: CARRIER SPACING FAULT
   RUNG wire#powerrail
      Contact( "reset" )
      Contact( "EMS".Carrier[31].SDC_OUT.Faults.CarrierSpacingFault )
      wire#w1
      Coil( "DB302_HMI_Faults".Carrier31_Faults_2.%X2 )
   END_RUNG
   RUNG wire#powerrail
      Contact( "DB302_HMI_Faults".Carrier31_Faults_2.%X2 )
      I_Contact( "EMS_Fault_Reset" )
   END_RUNG wire#w1
   // the same network as SCL:
   "DB302_HMI_Faults".Carrier31_Faults_2.%X2 := ("reset" AND "EMS".Carrier[31].SDC_OUT.Faults.CarrierSpacingFault) OR ("DB302_HMI_Faults".Carrier31_Faults_2.%X2 AND NOT "EMS_Fault_Reset");
END_REGION

REGION Network 36: DUPLICATE CARRIER NUMBER FAULT